screen "Last_1" 800x480, template "Main"
   TextField "Text field_1" at 220,5 size 368x47; Text 'Статистика весов 1'
   Button "HmiScreenItemData_1" at 10,425 size 159x47; TextOff 'Прошлый месяц'; TextOn 'Система'; PictureOn "Navigates to System screens for KTP700 Basic+ PN 14.0.1.0"; PictureOff "Navigates to System screens for KTP700 Basic+ PN 14.0.1.0"; Authorization "Admin"
   Button "HmiScreenItemData_4" at 565,425 size 159x47; TextOn 'О нас'; TextOff 'Текущий месяц'; PictureOn "Navigates to System screens for KTP700 Basic+ PN 14.0.1.0"; PictureOff "Navigates to System screens for KTP700 Basic+ PN 14.0.1.0"
      on Release: ActivateScreen("Mass_1", 0)
   TextField "Text field_4" at 12,61 size 61x23; Text 'День 1'
   TextField "Text field_5" at 12,97 size 61x23; Text 'День 2'
   TextField "Text field_6" at 12,134 size 61x23; Text 'День 3'
   TextField "Text field_7" at 12,170 size 61x23; Text 'День 4'
   TextField "Text field_8" at 12,207 size 61x23; Text 'День 5'
   TextField "Text field_9" at 12,243 size 61x23; Text 'День 6'
   TextField "Text field_10" at 12,280 size 61x23; Text 'День 7'
   TextField "Text field_11" at 12,316 size 61x23; Text 'День 8'
   TextField "Text field_12" at 12,353 size 61x23; Text 'День 9'
   TextField "Text field_13" at 12,390 size 71x23; Text 'День 10'
   IOField "I/O field_8" at 90,59 size 80x27; Authorization "Operator"; FormatPattern 999999.9
      ProcessValue <- "Statistics_DB_Last_M_1{1}"
   IOField "I/O field_3" at 90,95 size 80x27; Authorization "Operator"; FormatPattern 999999.9
      ProcessValue <- "Statistics_DB_Last_M_1{2}"
   IOField "I/O field_4" at 90,132 size 80x27; Authorization "Operator"; FormatPattern 999999.9
      ProcessValue <- "Statistics_DB_Last_M_1{3}"
   IOField "I/O field_5" at 90,168 size 80x27; Authorization "Operator"; FormatPattern 999999.9
      ProcessValue <- "Statistics_DB_Last_M_1{4}"
   IOField "I/O field_6" at 90,205 size 80x27; Authorization "Operator"; FormatPattern 999999.9
      ProcessValue <- "Statistics_DB_Last_M_1{5}"
   IOField "I/O field_7" at 90,241 size 80x27; Authorization "Operator"; FormatPattern 999999.9
      ProcessValue <- "Statistics_DB_Last_M_1{6}"
   IOField "I/O field_9" at 90,278 size 80x27; Authorization "Operator"; FormatPattern 999999.9
      ProcessValue <- "Statistics_DB_Last_M_1{7}"
   IOField "I/O field_10" at 90,314 size 80x27; Authorization "Operator"; FormatPattern 999999.9
      ProcessValue <- "Statistics_DB_Last_M_1{8}"
   IOField "I/O field_11" at 90,351 size 80x27; Authorization "Operator"; FormatPattern 999999.9
      ProcessValue <- "Statistics_DB_Last_M_1{9}"
   IOField "I/O field_12" at 90,388 size 80x27; Authorization "Operator"; FormatPattern 999999.9
      ProcessValue <- "Statistics_DB_Last_M_1{10}"
   IOField "I/O field_13" at 565,316 size 159x30; FormatPattern 99999.9
      Appearance <- "DIx_DB_Mass_1_Signal"
      ProcessValue <- "Statistics_DB_Last_Month_1"
   TextField "Text field_14" at 595,284 size 100x27; Text 'За месяц:'
   TextField "Text field_15" at 611,359 size 67x27; Text 'Всего:'
   IOField "I/O field_14" at 565,387 size 159x30; FormatPattern 9999999.9
      ProcessValue <- "Statistics_DB_All_1"
      Appearance <- "DIx_DB_Mass_1_Signal"
   TextField "Text field_16" at 202,62 size 71x23; Text 'День 11'
   TextField "Text field_18" at 202,98 size 71x23; Text 'День 12'
   TextField "Text field_19" at 202,135 size 71x23; Text 'День 13'
   TextField "Text field_20" at 202,171 size 71x23; Text 'День 14'
   TextField "Text field_21" at 202,208 size 71x23; Text 'День 15'
   TextField "Text field_22" at 202,244 size 71x23; Text 'День 16'
   TextField "Text field_23" at 202,281 size 71x23; Text 'День 17'
   TextField "Text field_24" at 202,317 size 71x23; Text 'День 18'
   TextField "Text field_25" at 202,354 size 71x23; Text 'День 19'
   TextField "Text field_26" at 202,391 size 71x23; Text 'День 20'
   IOField "I/O field_15" at 280,60 size 80x27; Authorization "Operator"; FormatPattern 999999.9
      ProcessValue <- "Statistics_DB_Last_M_1{11}"
   IOField "I/O field_16" at 280,96 size 80x27; Authorization "Operator"; FormatPattern 999999.9
      ProcessValue <- "Statistics_DB_Last_M_1{12}"
   IOField "I/O field_17" at 280,133 size 80x27; Authorization "Operator"; FormatPattern 999999.9
      ProcessValue <- "Statistics_DB_Last_M_1{13}"
   IOField "I/O field_18" at 280,169 size 80x27; Authorization "Operator"; FormatPattern 999999.9
      ProcessValue <- "Statistics_DB_Last_M_1{14}"
   IOField "I/O field_19" at 280,206 size 80x27; Authorization "Operator"; FormatPattern 999999.9
      ProcessValue <- "Statistics_DB_Last_M_1{15}"
   IOField "I/O field_20" at 280,242 size 80x27; Authorization "Operator"; FormatPattern 999999.9
      ProcessValue <- "Statistics_DB_Last_M_1{16}"
   IOField "I/O field_21" at 280,279 size 80x27; Authorization "Operator"; FormatPattern 999999.9
      ProcessValue <- "Statistics_DB_Last_M_1{17}"
   IOField "I/O field_22" at 280,315 size 80x27; Authorization "Operator"; FormatPattern 999999.9
      ProcessValue <- "Statistics_DB_Last_M_1{18}"
   IOField "I/O field_23" at 280,352 size 80x27; Authorization "Operator"; FormatPattern 999999.9
      ProcessValue <- "Statistics_DB_Last_M_1{19}"
   IOField "I/O field_24" at 280,389 size 80x27; Authorization "Operator"; FormatPattern 999999.9
      ProcessValue <- "Statistics_DB_Last_M_1{20}"
   TextField "Text field_27" at 392,63 size 71x23; Text 'День 21'
   TextField "Text field_28" at 392,99 size 71x23; Text 'День 22'
   TextField "Text field_29" at 392,136 size 71x23; Text 'День 23'
   TextField "Text field_30" at 392,172 size 71x23; Text 'День 24'
   TextField "Text field_31" at 392,209 size 71x23; Text 'День 25'
   TextField "Text field_32" at 392,245 size 71x23; Text 'День 26'
   TextField "Text field_33" at 392,282 size 71x23; Text 'День 27'
   TextField "Text field_34" at 392,318 size 71x23; Text 'День 28'
   TextField "Text field_35" at 392,355 size 71x23; Text 'День 29'
   TextField "Text field_36" at 392,392 size 71x23; Text 'День 30'
   IOField "I/O field_25" at 470,61 size 80x27; Authorization "Operator"; FormatPattern 999999.9
      ProcessValue <- "Statistics_DB_Last_M_1{21}"
   IOField "I/O field_26" at 470,97 size 80x27; Authorization "Operator"; FormatPattern 999999.9
      ProcessValue <- "Statistics_DB_Last_M_1{22}"
   IOField "I/O field_27" at 470,134 size 80x27; Authorization "Operator"; FormatPattern 999999.9
      ProcessValue <- "Statistics_DB_Last_M_1{23}"
   IOField "I/O field_28" at 470,170 size 80x27; Authorization "Operator"; FormatPattern 999999.9
      ProcessValue <- "Statistics_DB_Last_M_1{24}"
   IOField "I/O field_29" at 470,207 size 80x27; Authorization "Operator"; FormatPattern 999999.9
      ProcessValue <- "Statistics_DB_Last_M_1{25}"
   IOField "I/O field_30" at 470,243 size 80x27; Authorization "Operator"; FormatPattern 999999.9
      ProcessValue <- "Statistics_DB_Last_M_1{26}"
   IOField "I/O field_31" at 470,280 size 80x27; Authorization "Operator"; FormatPattern 999999.9
      ProcessValue <- "Statistics_DB_Last_M_1{27}"
   IOField "I/O field_32" at 470,316 size 80x27; Authorization "Operator"; FormatPattern 999999.9
      ProcessValue <- "Statistics_DB_Last_M_1{28}"
   IOField "I/O field_33" at 470,353 size 80x27; Authorization "Operator"; FormatPattern 999999.9
      ProcessValue <- "Statistics_DB_Last_M_1{29}"
   IOField "I/O field_34" at 470,390 size 80x27; Authorization "Operator"; FormatPattern 999999.9
      ProcessValue <- "Statistics_DB_Last_M_1{30}"
   TextField "Text field_37" at 563,64 size 71x23; Text 'День 31'
   IOField "I/O field_35" at 644,62 size 80x27; Authorization "Operator"; FormatPattern 999999.9
      ProcessValue <- "Statistics_DB_Last_M_1{31}"

screen "Last_2" 800x480, template "Main"
   TextField "Text field_1" at 220,5 size 368x47; Text 'Статистика весов 2'
   Button "HmiScreenItemData_1" at 10,425 size 159x47; TextOff 'Прошлый месяц'; TextOn 'Система'; Authorization "Admin"; PictureOff "Navigates to System screens for KTP700 Basic+ PN 14.0.1.0"; PictureOn "Navigates to System screens for KTP700 Basic+ PN 14.0.1.0"
   Button "HmiScreenItemData_4" at 565,425 size 159x47; TextOn 'О нас'; TextOff 'Текущий месяц'; PictureOn "Navigates to System screens for KTP700 Basic+ PN 14.0.1.0"; PictureOff "Navigates to System screens for KTP700 Basic+ PN 14.0.1.0"
      on Release: ActivateScreen("Mass_2", 0)
   TextField "Text field_5" at 12,61 size 61x23; Text 'День 1'
   TextField "Text field_6" at 12,97 size 61x23; Text 'День 2'
   TextField "Text field_7" at 12,134 size 61x23; Text 'День 3'
   TextField "Text field_8" at 12,170 size 61x23; Text 'День 4'
   TextField "Text field_9" at 12,207 size 61x23; Text 'День 5'
   TextField "Text field_10" at 12,243 size 61x23; Text 'День 6'
   TextField "Text field_11" at 12,280 size 61x23; Text 'День 7'
   TextField "Text field_12" at 12,316 size 61x23; Text 'День 8'
   TextField "Text field_13" at 12,353 size 61x23; Text 'День 9'
   TextField "Text field_14" at 12,390 size 71x23; Text 'День 10'
   IOField "I/O field_8" at 90,59 size 80x27; Authorization "Operator"; FormatPattern 999999.9
      ProcessValue <- "Statistics_DB_Last_M_2{1}"
   IOField "I/O field_3" at 90,95 size 80x27; Authorization "Operator"; FormatPattern 999999.9
      ProcessValue <- "Statistics_DB_Last_M_2{2}"
   IOField "I/O field_4" at 90,132 size 80x27; Authorization "Operator"; FormatPattern 999999.9
      ProcessValue <- "Statistics_DB_Last_M_2{3}"
   IOField "I/O field_5" at 90,168 size 80x27; Authorization "Operator"; FormatPattern 999999.9
      ProcessValue <- "Statistics_DB_Last_M_2{4}"
   IOField "I/O field_6" at 90,205 size 80x27; Authorization "Operator"; FormatPattern 999999.9
      ProcessValue <- "Statistics_DB_Last_M_2{5}"
   IOField "I/O field_7" at 90,241 size 80x27; Authorization "Operator"; FormatPattern 999999.9
      ProcessValue <- "Statistics_DB_Last_M_2{6}"
   IOField "I/O field_9" at 90,278 size 80x27; Authorization "Operator"; FormatPattern 999999.9
      ProcessValue <- "Statistics_DB_Last_M_2{7}"
   IOField "I/O field_10" at 90,314 size 80x27; Authorization "Operator"; FormatPattern 999999.9
      ProcessValue <- "Statistics_DB_Last_M_2{8}"
   IOField "I/O field_11" at 90,351 size 80x27; Authorization "Operator"; FormatPattern 999999.9
      ProcessValue <- "Statistics_DB_Last_M_2{9}"
   IOField "I/O field_12" at 90,388 size 80x27; Authorization "Operator"; FormatPattern 999999.9
      ProcessValue <- "Statistics_DB_Last_M_2{10}"
   IOField "I/O field_13" at 565,316 size 159x30; FormatPattern 99999.9
      Appearance <- "DIx_DB_Mass_2_Signal"
      ProcessValue <- "Statistics_DB_Last_Month_2"
   TextField "Text field_15" at 595,284 size 100x27; Text 'За месяц:'
   TextField "Text field_16" at 611,359 size 67x27; Text 'Всего:'
   IOField "I/O field_14" at 565,387 size 159x30; FormatPattern 9999999.9
      ProcessValue <- "Statistics_DB_All_2"
      Appearance <- "DIx_DB_Mass_2_Signal"
   TextField "Text field_18" at 202,62 size 71x23; Text 'День 11'
   TextField "Text field_19" at 202,98 size 71x23; Text 'День 12'
   TextField "Text field_20" at 202,135 size 71x23; Text 'День 13'
   TextField "Text field_21" at 202,171 size 71x23; Text 'День 14'
   TextField "Text field_22" at 202,208 size 71x23; Text 'День 15'
   TextField "Text field_23" at 202,244 size 71x23; Text 'День 16'
   TextField "Text field_24" at 202,281 size 71x23; Text 'День 17'
   TextField "Text field_25" at 202,317 size 71x23; Text 'День 18'
   TextField "Text field_26" at 202,354 size 71x23; Text 'День 19'
   TextField "Text field_27" at 202,391 size 71x23; Text 'День 20'
   IOField "I/O field_15" at 280,60 size 80x27; Authorization "Operator"; FormatPattern 999999.9
      ProcessValue <- "Statistics_DB_Last_M_2{11}"
   IOField "I/O field_16" at 280,96 size 80x27; Authorization "Operator"; FormatPattern 999999.9
      ProcessValue <- "Statistics_DB_Last_M_2{12}"
   IOField "I/O field_17" at 280,133 size 80x27; Authorization "Operator"; FormatPattern 999999.9
      ProcessValue <- "Statistics_DB_Last_M_2{13}"
   IOField "I/O field_18" at 280,169 size 80x27; Authorization "Operator"; FormatPattern 999999.9
      ProcessValue <- "Statistics_DB_Last_M_2{14}"
   IOField "I/O field_19" at 280,206 size 80x27; Authorization "Operator"; FormatPattern 999999.9
      ProcessValue <- "Statistics_DB_Last_M_2{15}"
   IOField "I/O field_20" at 280,242 size 80x27; Authorization "Operator"; FormatPattern 999999.9
      ProcessValue <- "Statistics_DB_Last_M_2{16}"
   IOField "I/O field_21" at 280,279 size 80x27; Authorization "Operator"; FormatPattern 999999.9
      ProcessValue <- "Statistics_DB_Last_M_2{17}"
   IOField "I/O field_22" at 280,315 size 80x27; Authorization "Operator"; FormatPattern 999999.9
      ProcessValue <- "Statistics_DB_Last_M_2{18}"
   IOField "I/O field_23" at 280,352 size 80x27; Authorization "Operator"; FormatPattern 999999.9
      ProcessValue <- "Statistics_DB_Last_M_2{19}"
   IOField "I/O field_24" at 280,389 size 80x27; Authorization "Operator"; FormatPattern 999999.9
      ProcessValue <- "Statistics_DB_Last_M_2{20}"
   TextField "Text field_28" at 392,63 size 71x23; Text 'День 21'
   TextField "Text field_29" at 392,99 size 71x23; Text 'День 22'
   TextField "Text field_30" at 392,136 size 71x23; Text 'День 23'
   TextField "Text field_31" at 392,172 size 71x23; Text 'День 24'
   TextField "Text field_32" at 392,209 size 71x23; Text 'День 25'
   TextField "Text field_33" at 392,245 size 71x23; Text 'День 26'
   TextField "Text field_34" at 392,282 size 71x23; Text 'День 27'
   TextField "Text field_35" at 392,318 size 71x23; Text 'День 28'
   TextField "Text field_36" at 392,355 size 71x23; Text 'День 29'
   TextField "Text field_37" at 392,392 size 71x23; Text 'День 30'
   IOField "I/O field_25" at 470,61 size 80x27; Authorization "Operator"; FormatPattern 999999.9
      ProcessValue <- "Statistics_DB_Last_M_2{21}"
   IOField "I/O field_26" at 470,97 size 80x27; Authorization "Operator"; FormatPattern 999999.9
      ProcessValue <- "Statistics_DB_Last_M_2{22}"
   IOField "I/O field_27" at 470,134 size 80x27; Authorization "Operator"; FormatPattern 999999.9
      ProcessValue <- "Statistics_DB_Last_M_2{23}"
   IOField "I/O field_28" at 470,170 size 80x27; Authorization "Operator"; FormatPattern 999999.9
      ProcessValue <- "Statistics_DB_Last_M_2{24}"
   IOField "I/O field_29" at 470,207 size 80x27; Authorization "Operator"; FormatPattern 999999.9
      ProcessValue <- "Statistics_DB_Last_M_2{25}"
   IOField "I/O field_30" at 470,243 size 80x27; Authorization "Operator"; FormatPattern 999999.9
      ProcessValue <- "Statistics_DB_Last_M_2{26}"
   IOField "I/O field_31" at 470,280 size 80x27; Authorization "Operator"; FormatPattern 999999.9
      ProcessValue <- "Statistics_DB_Last_M_2{27}"
   IOField "I/O field_32" at 470,316 size 80x27; Authorization "Operator"; FormatPattern 999999.9
      ProcessValue <- "Statistics_DB_Last_M_2{28}"
   IOField "I/O field_33" at 470,353 size 80x27; Authorization "Operator"; FormatPattern 999999.9
      ProcessValue <- "Statistics_DB_Last_M_2{29}"
   IOField "I/O field_34" at 470,390 size 80x27; Authorization "Operator"; FormatPattern 999999.9
      ProcessValue <- "Statistics_DB_Last_M_2{30}"
   TextField "Text field_38" at 563,64 size 71x23; Text 'День 31'
   IOField "I/O field_35" at 644,62 size 80x27; Authorization "Operator"; FormatPattern 999999.9
      ProcessValue <- "Statistics_DB_Last_M_2{31}"

screen "PID_settings" 800x480, template "Main"
   TextField "Text field_1" at 133,9 size 84x22; Text 'ПИД: M1'
   Button "Button_14" at 157,37 size 68x28; TextOff 'Hand'
      on Click: InvertBit("PID_M1_Hand")
      Appearance <- "PID_M1_Hand"
   IOField "I/O field_29" at 230,37 size 78x28; FormatPattern s9999.9
      ProcessValue <- "PID_M1_HandValue"
   Button "Button_1" at 314,37 size 68x28; TextOff 'Reset'
      on Click: InvertBit("PID_M1_Reset")
      Appearance <- "PID_M1_Reset"
   TextField "Text field_25" at 131,93 size 19x28; Text 'K'
   TextField "Text field_26" at 131,124 size 23x28; Text 'Ti'
   TextField "Text field_27" at 131,155 size 30x28; Text 'Td'
   IOField "I/O field_32" at 165,91 size 60x30; FormatPattern 99999
      ProcessValue <- "PID_M1_SP_P"
   IOField "I/O field_33" at 165,122 size 60x30; FormatPattern 99999
      ProcessValue <- "PID_M1_SP_Ti"
   IOField "I/O field_34" at 165,153 size 60x30; FormatPattern 99999
      ProcessValue <- "PID_M1_SP_Td"
   TextField "Text field_2" at 131,202 size 73x22; Text 'Уставка:'
   TextField "Text field_4" at 131,223 size 67x22; Text 'Датчик:'
   IOField "I/O field_1" at 309,201 size 58x21; FormatPattern 99999
      ProcessValue <- "PID_M1_Max_SP"
   IOField "I/O field_2" at 236,202 size 58x21; FormatPattern 99999
      ProcessValue <- "PID_M1_Min_SP"
   IOField "I/O field_3" at 309,222 size 58x21; FormatPattern s99999
      ProcessValue <- "PID_M1_Max_in"
   IOField "I/O field_4" at 236,223 size 58x21; FormatPattern s99999
      ProcessValue <- "PID_M1_Min_in"
   TextField "Text field_8" at 131,244 size 62x22; Text 'Выход:'
   IOField "I/O field_5" at 309,243 size 58x21; FormatPattern 99999
      ProcessValue <- "PID_M1_Max_out"
   IOField "I/O field_6" at 236,244 size 58x21; FormatPattern 99999
      ProcessValue <- "PID_M1_Min_out"
   TextField "Text field_12" at 320,177 size 36x22; Text 'Max'
   TextField "Text field_14" at 249,178 size 32x22; Text 'Min'
   TextField "Text field_3" at 257,91 size 31x28; Text 'SP'
   IOField "I/O field_9" at 323,89 size 60x30; FormatPattern 99999
      ProcessValue <- "PID_M1_SP"
   TextField "Text field_7" at 257,122 size 62x28; Text 'Value'
   IOField "I/O field_10" at 323,120 size 60x30; FormatPattern 99999
      ProcessValue <- "PID_M1_Value"
   Button "Button_2" at 346,281 size 58x28; TextOff 'Inv'
      on Click: InvertBit("PID_M1_Invert")
      Appearance <- "PID_M1_Invert"
   TextField "Text field_28" at 130,280 size 109x22; Text 'Время цикла:'
   IOField "I/O field_35" at 280,281 size 58x21; FormatPattern s99999
      ProcessValue <- "PID_M1_SP_Cycle"
   TextField "Text field_10" at 130,302 size 116x22; Text 'Мертвая зона:'
   TextField "Text field_11" at 130,353 size 132x22; Text 'Входной сигнал:'
   IOField "I/O field_7" at 280,303 size 58x21; FormatPattern s99999
      ProcessValue <- "PID_M1_DeadBand"
   IOField "I/O field_8" at 346,354 size 58x21; FormatPattern s99999
      ProcessValue <- "PID_M1_Converter_Max_In"
   IOField "I/O field_11" at 278,354 size 58x21; FormatPattern s99999
      ProcessValue <- "PID_M1_Converter_Min_In"
   TextField "Text field_13" at 130,375 size 145x22; Text 'Выходной сигнал:'
   IOField "I/O field_12" at 346,376 size 58x21; FormatPattern s99999
      ProcessValue <- "PID_M1_Converter_Max_Out"
   IOField "I/O field_13" at 278,376 size 58x21; FormatPattern s99999
      ProcessValue <- "PID_M1_Converter_Min_Out"
   TextField "Text field_5" at 357,332 size 36x22; Text 'Max'
   TextField "Text field_6" at 278,332 size 32x22; Text 'Min'
   TextField "Text field_9" at 443,8 size 84x22; Text 'ПИД: M2'
   Button "Button_9" at 467,36 size 68x28; TextOff 'Hand'
      on Click: InvertBit("PID_M2_Hand")
      Appearance <- "PID_M2_Hand"
   IOField "I/O field_14" at 540,36 size 78x28; FormatPattern s9999.9
      ProcessValue <- "PID_M2_HandValue"
   Button "Button_10" at 624,36 size 68x28; TextOff 'Reset'
      on Click: InvertBit("PID_M2_Reset")
      Appearance <- "PID_M2_Reset"
   TextField "Text field_15" at 441,92 size 19x28; Text 'K'
   TextField "Text field_16" at 441,123 size 23x28; Text 'Ti'
   TextField "Text field_17" at 441,154 size 30x28; Text 'Td'
   IOField "I/O field_15" at 475,90 size 60x30; FormatPattern 99999
      ProcessValue <- "PID_M2_SP_P"
   IOField "I/O field_16" at 475,121 size 60x30; FormatPattern 99999
      ProcessValue <- "PID_M2_SP_Ti"
   IOField "I/O field_17" at 475,152 size 60x30; FormatPattern 99999
      ProcessValue <- "PID_M2_SP_Td"
   TextField "Text field_18" at 441,201 size 73x22; Text 'Уставка:'
   TextField "Text field_19" at 441,222 size 67x22; Text 'Датчик:'
   IOField "I/O field_18" at 619,200 size 58x21; FormatPattern 99999
      ProcessValue <- "PID_M2_Max_SP"
   IOField "I/O field_19" at 546,201 size 58x21; FormatPattern 99999
      ProcessValue <- "PID_M2_Min_SP"
   IOField "I/O field_20" at 619,221 size 58x21; FormatPattern s99999
      ProcessValue <- "PID_M2_Max_in"
   IOField "I/O field_21" at 546,222 size 58x21; FormatPattern s99999
      ProcessValue <- "PID_M2_Min_in"
   TextField "Text field_20" at 441,243 size 62x22; Text 'Выход:'
   IOField "I/O field_22" at 619,242 size 58x21; FormatPattern 99999
      ProcessValue <- "PID_M2_Max_out"
   IOField "I/O field_23" at 546,243 size 58x21; FormatPattern 99999
      ProcessValue <- "PID_M2_Min_out"
   TextField "Text field_21" at 630,176 size 36x22; Text 'Max'
   TextField "Text field_22" at 559,177 size 32x22; Text 'Min'
   TextField "Text field_23" at 567,90 size 31x28; Text 'SP'
   IOField "I/O field_24" at 633,88 size 60x30; FormatPattern 99999
      ProcessValue <- "PID_M2_SP"
   TextField "Text field_24" at 567,121 size 62x28; Text 'Value'
   IOField "I/O field_25" at 633,119 size 60x30; FormatPattern 99999
      ProcessValue <- "PID_M2_Value"
   Button "Button_11" at 656,280 size 58x28; TextOff 'Inv'
      on Click: InvertBit("PID_M2_Invert")
      Appearance <- "PID_M2_Invert"
   TextField "Text field_29" at 440,279 size 109x22; Text 'Время цикла:'
   IOField "I/O field_26" at 590,280 size 58x21; FormatPattern s99999
      ProcessValue <- "PID_M2_SP_Cycle"
   TextField "Text field_30" at 440,301 size 116x22; Text 'Мертвая зона:'
   TextField "Text field_31" at 440,352 size 132x22; Text 'Входной сигнал:'
   IOField "I/O field_27" at 590,302 size 58x21; FormatPattern s99999
      ProcessValue <- "PID_M2_DeadBand"
   IOField "I/O field_28" at 656,353 size 58x21; FormatPattern s99999
      ProcessValue <- "PID_M2_Converter_Max_In"
   IOField "I/O field_30" at 588,353 size 58x21; FormatPattern s99999
      ProcessValue <- "PID_M2_Converter_Min_In"
   TextField "Text field_32" at 440,374 size 145x22; Text 'Выходной сигнал:'
   IOField "I/O field_31" at 656,375 size 58x21; FormatPattern s99999
      ProcessValue <- "PID_M2_Converter_Max_Out"
   IOField "I/O field_36" at 588,375 size 58x21; FormatPattern s99999
      ProcessValue <- "PID_M2_Converter_Min_Out"
   TextField "Text field_33" at 667,331 size 36x22; Text 'Max'
   TextField "Text field_34" at 588,331 size 32x22; Text 'Min'
   Button "Button_3" at 7,5 size 96x32; TextOff 'Насосы'; Authorization "Admin"
      on Release: ActivateScreen("Dos", 0); SetTag("settings", 1)
      Appearance <- "settings"
   Button "Button_4" at 7,51 size 96x32; TextOff 'Расход-1'; Authorization "Admin"
      on Release: ActivateScreen("Flow", 0); SetTag("settings", 2)
      Appearance <- "settings"
   Button "Button_5" at 7,140 size 96x32; TextOff 'Мутность'; Authorization "Admin"
      on Release: ActivateScreen("Trans", 0); SetTag("settings", 4)
      Appearance <- "settings"
   Button "Button_6" at 7,184 size 96x32; TextOff 'DI'; Authorization "Admin"
      on Release: ActivateScreen("DI", 0); SetTag("settings", 5)
      Appearance <- "settings"
   Button "Button_7" at 7,229 size 96x32; TextOff 'DO'; Authorization "Admin"
      on Release: ActivateScreen("DO", 0); SetTag("settings", 6)
      Appearance <- "settings"
   Button "Button_8" at 7,274 size 96x32; TextOff 'PID'; Authorization "Admin"
      on Release: ActivateScreen("PID_settings", 0); SetTag("settings", 7)
      Appearance <- "settings"
   Button "Button_15" at 7,95 size 96x32; TextOff 'Расход-2'; Authorization "Admin"
      on Release: ActivateScreen("Flow_1", 0); SetTag("settings", 3)
      Appearance <- "settings"

screen "Flow_1" 800x480, template "Main"
   TextField "Text field_2" at 210,15 size 67x22; Text 'Датчик:'
   TextField "Text field_4" at 273,15 size 113x22; Text 'Расходомер 3'
   TextField "Text field_7" at 390,18 size 43x22; Text 'вход'
   TextField "Text field_8" at 390,43 size 56x22; Text 'выход'
   IOField "I/O field_1" at 452,19 size 102x26; FormatPattern s99999.99
      ProcessValue <- "AIx_DB_Flow_3_Converter_Min_In"
   IOField "I/O field_2" at 452,41 size 102x26; FormatPattern s99999.99
      ProcessValue <- "AIx_DB_Flow_3_Converter_Min_Out"
   IOField "I/O field_3" at 551,19 size 102x26; FormatPattern s99999.99
      ProcessValue <- "AIx_DB_Flow_3_Converter_Max_In"
   IOField "I/O field_4" at 551,41 size 102x26; FormatPattern s99999.99
      ProcessValue <- "AIx_DB_Flow_3_Converter_Max_Out"
   TextField "Text field_9" at 389,68 size 101x22; Text 'Фильтрация'
   TextField "Text field_10" at 390,96 size 36x22; Text 'RTD'
   Button "Button_7" at 489,71 size 20x20; TextOff 'Text'; PictureList "ok"
      on Click: InvertBit("AIx_DB_Flow_3_Use_Filter")
      ProcessValue <- "AIx_DB_Flow_3_Use_Filter"
   Button "Button_8" at 489,96 size 20x20; TextOff 'Text'; PictureList "ok"
      on Click: InvertBit("AIx_DB_Flow_3_Use_RTD")
      ProcessValue <- "AIx_DB_Flow_3_Use_RTD"
   IOField "I/O field_5" at 516,68 size 65x25; FormatPattern 999
      ProcessValue <- "AIx_DB_Flow_3_Filter_SP"
   IOField "I/O field_6" at 516,93 size 65x25; FormatPattern 999
      ProcessValue <- "AIx_DB_Flow_3_RTD_c"
   TextField "Text field_11" at 210,36 size 79x22; Text 'Поправка'
   IOField "I/O field_7" at 293,36 size 78x23; FormatPattern s999.9
      ProcessValue <- "AIx_DB_Flow_3_Calibration"
   Button "Button_9" at 396,176 size 248x28; TextOff 'Use'
      on Click: InvertBit("AIx_DB_Flow_3_CMD_Start_A")
      Appearance <- "AIx_DB_Flow_3_CMD_Start_A"
   Button "Button_10" at 213,66 size 68x28; TextOff 'Hand'
      on Click: InvertBit("AIx_DB_Flow_3_CMD_Hand")
      Appearance <- "AIx_DB_Flow_3_CMD_Hand"
   IOField "I/O field_8" at 293,66 size 78x28; FormatPattern s9999.9
      ProcessValue <- "AIx_DB_Flow_3_Result"
   TextField "Text field_12" at 436,123 size 27x22; Text 'NC'
   TextField "Text field_13" at 437,143 size 25x22; Text 'SC'
   TextField "Text field_14" at 210,125 size 27x22; Text 'HH'
   TextField "Text field_15" at 216,145 size 16x22; Text 'H'
   TextField "Text field_16" at 217,165 size 14x22; Text 'L'
   TextField "Text field_17" at 212,186 size 23x22; Text 'LL'
   IOField "I/O field_11" at 472,123 size 58x21; FormatPattern s99999
      ProcessValue <- "AIx_DB_Flow_3_SP_NC"
   IOField "I/O field_12" at 472,143 size 58x21; FormatPattern s99999
      ProcessValue <- "AIx_DB_Flow_3_SP_SC"
   IOField "I/O field_13" at 246,125 size 58x21; FormatPattern 99999
      ProcessValue <- "AIx_DB_Flow_3_SP_HH"
   IOField "I/O field_14" at 246,145 size 58x21; FormatPattern 99999
      ProcessValue <- "AIx_DB_Flow_3_SP_H"
   IOField "I/O field_15" at 246,165 size 58x21; FormatPattern s99999
      ProcessValue <- "AIx_DB_Flow_3_SP_L"
   IOField "I/O field_16" at 246,185 size 58x21; FormatPattern s99999
      ProcessValue <- "AIx_DB_Flow_3_SP_LL"
   IOField "I/O field_17" at 546,123 size 58x21; FormatPattern 999
      ProcessValue <- "AIx_DB_Flow_3_Timers_NC_SP"
   IOField "I/O field_18" at 546,143 size 58x21; FormatPattern 999
      ProcessValue <- "AIx_DB_Flow_3_Timers_SC_SP"
   IOField "I/O field_19" at 320,125 size 58x21; FormatPattern 999
      ProcessValue <- "AIx_DB_Flow_3_Timers_HH_SP"
   IOField "I/O field_20" at 320,145 size 58x21; FormatPattern 999
      ProcessValue <- "AIx_DB_Flow_3_Timers_H_SP"
   IOField "I/O field_21" at 320,165 size 58x21; FormatPattern 999
      ProcessValue <- "AIx_DB_Flow_3_Timers_L_SP"
   IOField "I/O field_22" at 320,185 size 58x21; FormatPattern 999
      ProcessValue <- "AIx_DB_Flow_3_Timers_LL_SP"
   IOField "I/O field_23" at 582,93 size 65x25; FormatPattern s99999
      ProcessValue <- "AIx_DB_Flow_3_Signal"
   TextField "Text field_18" at 210,97 size 68x22; Text 'Уставка'
   TextField "Text field_19" at 299,97 size 79x22; Text 'Время (с)'
   TextField "Text field_1" at 214,248 size 67x22; Text 'Датчик:'
   TextField "Text field_3" at 277,248 size 113x22; Text 'Расходомер 4'
   TextField "Text field_5" at 394,251 size 43x22; Text 'вход'
   TextField "Text field_6" at 394,276 size 56x22; Text 'выход'
   IOField "I/O field_9" at 456,252 size 102x26; FormatPattern s99999.99
      ProcessValue <- "AIx_DB_Flow_4_Converter_Min_In"
   IOField "I/O field_10" at 456,274 size 102x26; FormatPattern s99999.99
      ProcessValue <- "AIx_DB_Flow_4_Converter_Min_Out"
   IOField "I/O field_24" at 555,252 size 102x26; FormatPattern s99999.99
      ProcessValue <- "AIx_DB_Flow_4_Converter_Max_In"
   IOField "I/O field_25" at 555,274 size 102x26; FormatPattern s99999.99
      ProcessValue <- "AIx_DB_Flow_4_Converter_Max_Out"
   TextField "Text field_20" at 393,301 size 101x22; Text 'Фильтрация'
   TextField "Text field_21" at 394,329 size 36x22; Text 'RTD'
   Button "Button_11" at 493,304 size 20x20; TextOff 'Text'; PictureList "ok"
      on Click: InvertBit("AIx_DB_Flow_4_Use_Filter")
      ProcessValue <- "AIx_DB_Flow_4_Use_Filter"
   Button "Button_12" at 493,329 size 20x20; TextOff 'Text'; PictureList "ok"
      on Click: InvertBit("AIx_DB_Flow_4_Use_RTD")
      ProcessValue <- "AIx_DB_Flow_4_Use_RTD"
   IOField "I/O field_26" at 520,301 size 65x25; FormatPattern 999
      ProcessValue <- "AIx_DB_Flow_4_Filter_SP"
   IOField "I/O field_27" at 520,326 size 65x25; FormatPattern 999
      ProcessValue <- "AIx_DB_Flow_4_RTD_c"
   TextField "Text field_22" at 214,269 size 79x22; Text 'Поправка'
   IOField "I/O field_28" at 297,269 size 78x23; FormatPattern s999.9
      ProcessValue <- "AIx_DB_Flow_4_Calibration"
   Button "Button_13" at 400,409 size 248x28; TextOff 'Use'
      on Click: InvertBit("AIx_DB_Flow_4_CMD_Start_A")
      Appearance <- "AIx_DB_Flow_4_CMD_Start_A"
   Button "Button_14" at 217,299 size 68x28; TextOff 'Hand'
      on Click: InvertBit("AIx_DB_Flow_4_CMD_Hand")
      Appearance <- "AIx_DB_Flow_4_CMD_Hand"
   IOField "I/O field_29" at 297,299 size 78x28; FormatPattern s9999.9
      ProcessValue <- "AIx_DB_Flow_4_Result"
   TextField "Text field_23" at 440,356 size 27x22; Text 'NC'
   TextField "Text field_24" at 441,376 size 25x22; Text 'SC'
   TextField "Text field_25" at 214,358 size 27x22; Text 'HH'
   TextField "Text field_26" at 220,378 size 16x22; Text 'H'
   TextField "Text field_27" at 221,398 size 14x22; Text 'L'
   TextField "Text field_28" at 216,419 size 23x22; Text 'LL'
   IOField "I/O field_30" at 476,356 size 58x21; FormatPattern s99999
      ProcessValue <- "AIx_DB_Flow_4_SP_NC"